// TIA Portal project "THELMA3_200224" (V15.1) (continued)
VERSION : 0.1
   STRUCT
      RemoteAddress : String;
      NonMDR_LabelName : String;
      "Date" : String;
      "Time" : String;
      RData : Array[0..56] of Byte;
      RdataBatch : Array[0..56] of Byte;
      BatchOK : Bool;
      TimeOK : Bool;
      AlarmCheck : Bool;
      LabelOK : Bool;
      LED_State : USInt;
      TimeDateError : Bool;
      Initialization : Bool;
      OPC_Error : Bool;
      TCP_ComError : Bool;
      TCP_ComErrorBatch : Bool;
      ComErrorStatus : Byte;
      ComErrorStatusBatch : Byte;
   END_STRUCT;
END_TYPE

TYPE "typeLCom_Config"
VERSION : 0.1
   STRUCT
      connection : Struct
         interfaceID : Hw_Any := 64;
         connectionID : Conn_Any := W#16#0FFF;
         comService : USInt := 2;
         isClient : Bool := false;
         localPort : UInt := 3456;
         partnerPort : UInt := 3456;
         partnerIP : IP_V4;
         acceptUnknownPartner : Bool := true;
         lifeSignCycleTime : Time := T#1s;
      END_STRUCT;
      sender : Struct
         cycleTime : Time := T#1s;
         ackTimeout : Time := T#1s;
      END_STRUCT;
      timeSync : Struct
         usePartnerTimestamps : Bool := false;
         sendMode : USInt;
         cycleTime : Time := T#1h;
         sendAtTimeOfDay : Time_Of_Day :=  TOD#05:00:0.000;
      END_STRUCT;
   END_STRUCT;
END_TYPE

TYPE "typeLCom_Diagnostics"
VERSION : 0.1
   STRUCT
      localConfig : Struct
         connection : Struct
            interfaceID : Hw_Any := 0;
            connectionID : Conn_Any := W#16#0000;
            comService : USInt := 0;
            isClient : Bool := false;
            localPort : UInt := 0;
            localIP : IP_V4;
            partnerPort : UInt := 3456;
            partnerIP : IP_V4;
            acceptUnknownPartner : Bool := false;
            useLComProtocol : Bool := false;
            lifeSignCycleTime : Time := T#0ms;
         END_STRUCT;
         sender : Struct
            cycleTime : Time;
            ackTimeout : Time;
         END_STRUCT;
         timeSync : Struct
            usePartnerTimestamps : Bool := false;
            sendMode : USInt;
            cycleTime : Time := T#0ms;
            sendAtTimeOfDay : Time_Of_Day :=  TOD#00:00:0.000;
         END_STRUCT;
         sizeOfSendBuffer : UDInt;
         sizeOfReceiveBuffer : UDInt;
      END_STRUCT;
      partnerConfig : Struct
         connnection : Struct
            lifeSignCycleTime : Time := T#0ms;
         END_STRUCT;
         sender : Struct
            cycleTime : Time := T#0ms;
            ackTimeout : Time := T#0ms;
         END_STRUCT;
         timeSync : Struct
            usePartnerTimestamps : Bool := false;
            sendMode : USInt;
         END_STRUCT;
         sizeOfSendBuffer : UDInt;
         sizeOfReceiveBuffer : UDInt;
      END_STRUCT;
      statistics : Struct
         avgCallCycle : Real;
         avgReceiveMsgCycle : Real;
         maxReceiveMsgCycle : Time;
         LComProtocolUsed : Bool := false;
         activeLComVersion : USInt;
         avgMsgSendingTime : Real;
         maxMsgSendingTime : Time;
         avgMsgReceivingTime : Real;
         maxMsgReceivingTime : Time;
         numberOfSentMessages : UDInt;
         numberOfReceivedMessages : UDInt;
         totalAckTimeouts : UInt;
         totalSendCycleViolations : UInt;
         totalReceiveCycleViolations : UInt;
         totalReconnects : UInt;
         lastConnect : DTL;
         lastTimeSync : DTL;
      END_STRUCT;
      bufferIndex : USInt := 16#FF;
      buffer : Array[0..63] of Struct
         status : Word;
         timestamp : DTL;
         isActive : Bool;
         subFunctionErrorID : Word;
         additionalValue1 : Real;
         additionalValue2 : Real;
         additionalValue3 : Real;
         additionalValue4 : Time;
      END_STRUCT;
   END_STRUCT;
   // buffer[1].isActive := false;
   // buffer[0].isActive := false;
   // buffer[2].isActive := false;
   // buffer[3].isActive := false;
   // buffer[4].isActive := false;
   // buffer[5].isActive := false;
   // buffer[6].isActive := false;
   // buffer[7].isActive := false;
   // buffer[8].isActive := false;
   // buffer[9].isActive := false;
   // buffer[10].isActive := false;
   // buffer[11].isActive := false;
   // buffer[12].isActive := false;
   // buffer[13].isActive := false;
   // buffer[14].isActive := false;
   // buffer[15].isActive := false;
   // buffer[16].isActive := false;
   // buffer[17].isActive := false;
   // buffer[18].isActive := false;
   // buffer[19].isActive := false;
   // buffer[20].isActive := false;
   // buffer[21].isActive := false;
   // buffer[22].isActive := false;
   // buffer[23].isActive := false;
   // buffer[24].isActive := false;
   // buffer[25].isActive := false;
   // buffer[26].isActive := false;
   // buffer[27].isActive := false;
   // buffer[28].isActive := false;
   // buffer[29].isActive := false;
   // buffer[30].isActive := false;
   // buffer[31].isActive := false;
   // buffer[32].isActive := false;
   // buffer[33].isActive := false;
   // buffer[34].isActive := false;
   // buffer[35].isActive := false;
   // buffer[36].isActive := false;
   // buffer[37].isActive := false;
   // buffer[38].isActive := false;
   // buffer[39].isActive := false;
   // buffer[40].isActive := false;
   // buffer[41].isActive := false;
   // buffer[42].isActive := false;
   // buffer[43].isActive := false;
   // buffer[44].isActive := false;
   // buffer[45].isActive := false;
   // buffer[46].isActive := false;
   // buffer[47].isActive := false;
   // buffer[48].isActive := false;
   // buffer[49].isActive := false;
   // buffer[50].isActive := false;
   // buffer[51].isActive := false;
   // buffer[52].isActive := false;
   // buffer[53].isActive := false;
   // buffer[54].isActive := false;
   // buffer[55].isActive := false;
   // buffer[56].isActive := false;
   // buffer[57].isActive := false;
   // buffer[58].isActive := false;
   // buffer[59].isActive := false;
   // buffer[60].isActive := false;
   // buffer[61].isActive := false;
   // buffer[62].isActive := false;
   // buffer[63].isActive := false;
END_TYPE

DATA_BLOCK "Skuska"   // DB1
{ S7_Optimized_Access := 'TRUE' }
VERSION : 0.1
   VAR
      SkuskaString : String;
      Length : Int;
      SkuskaArray : Array[0..56] of Byte;
      SkuskaString2 : String;
      TestBits : Array[0..10] of Bool;
      RemoteAdress : String := '192.168.1.10:29043';
   END_VAR
BEGIN
END_DATA_BLOCK

DATA_BLOCK "OPC"   // DB2
{ S7_Optimized_Access := 'TRUE' }
VERSION : 0.1
   VAR RETAIN
      CON_Material : "UDT_CON_Comm";
      TRP_Material : "UDT_TRP_Comm";
   END_VAR
BEGIN
END_DATA_BLOCK

DATA_BLOCK "SeP"   // DB3
{ S7_Optimized_Access := 'TRUE' }
VERSION : 0.1
   VAR
      Material_1 : "UDT_Status";
      Material_2 : "UDT_Status";
   END_VAR
BEGIN
END_DATA_BLOCK

DATA_BLOCK "LatestReading"   // DB4
{ S7_Optimized_Access := 'FALSE' }
VERSION : 0.1
   VAR
      TRP : "UDT_LatestReading";
   END_VAR
BEGIN
END_DATA_BLOCK

DATA_BLOCK "Reader"   // DB5
{ S7_Optimized_Access := 'TRUE' }
VERSION : 0.1
   VAR
      TRP : "UDT_Reader";
   END_VAR
BEGIN
END_DATA_BLOCK

DATA_BLOCK "TRP_DB"   // DB6
{ S7_Optimized_Access := 'TRUE' }
VERSION : 0.1
// stored: InstanceOfName TRP
"TRP"
BEGIN
END_DATA_BLOCK

DATA_BLOCK "CON_DB"   // DB7
{ S7_Optimized_Access := 'TRUE' }
VERSION : 0.1
// stored: InstanceOfName CON
"CON"
BEGIN
END_DATA_BLOCK

DATA_BLOCK "LatestReading_1"   // DB8
{ S7_Optimized_Access := 'FALSE' }
VERSION : 0.1
   VAR
      TRP : "UDT_LatestReading";
   END_VAR
BEGIN
END_DATA_BLOCK

DATA_BLOCK "PrinterData"   // DB9
{ S7_Optimized_Access := 'TRUE' }
VERSION : 0.1
   VAR RETAIN
      TRP : Struct
         PrinterData : "UDT_Printer";
         PrinterStatus : "typeLCom_Diagnostics";
         PrinterConfig : "typeLCom_Config";
      END_STRUCT;
      CON : Struct
         PrinterBagConfigBatch : "typeLCom_Config";
         PrinterBagStatusBatch : "typeLCom_Diagnostics";
         PrinterBagConfig : "typeLCom_Config";
         PrinterBagStatus : "typeLCom_Diagnostics";
         PrinterBagData : "UDT_CON_Printer";
         PrinterSelection : Bool;
      END_STRUCT;
   END_VAR
BEGIN
   TRP.PrinterData.RemoteAddress := '10.212.77.75:9100';
END_DATA_BLOCK

DATA_BLOCK "SiteCom"   // DB10
{ S7_Optimized_Access := 'FALSE' }
AUTHOR : nlagela
VERSION : 0.1
   VAR
      Material_1 : "UDT_ComMaterialReading";
      Material_2 : "UDT_ComMaterialReading";
   END_VAR
BEGIN
END_DATA_BLOCK

DATA_BLOCK "LatestReadings"   // DB11
{ S7_Optimized_Access := 'FALSE' }
VERSION : 0.1
   VAR
      Material_1 : "UDT_LatestReadingBag";
      Material_2 : "UDT_LatestReadingBag";
   END_VAR
BEGIN
END_DATA_BLOCK

DATA_BLOCK "PlainHandle_DB"   // DB12
{ S7_Optimized_Access := 'TRUE' }
VERSION : 0.1
// stored: InstanceOfName PlainHandle
"PlainHandle"
BEGIN
END_DATA_BLOCK

DATA_BLOCK "d10_PlainComm"   // DB13
{ S7_Optimized_Access := 'TRUE' }
VERSION : 0.1
   VAR
      Data_device : Array[0..7] of Bool;
   END_VAR
   VAR RETAIN
      bag_dmc_code : String [10];
      box_dmc_code : String [10];
      article_num : String [12];
      total_in_bag : String [7];
      total_in_box : String [7];
      product_weight : String [10];
      line_number : String [5];
      order_num : String [12];
   END_VAR
   VAR
      xPresetDataBagSent : Bool;
      xPresetDataBoxSent : Bool;
   END_VAR
BEGIN
END_DATA_BLOCK

DATA_BLOCK "d10_Data"   // DB14
{ S7_Optimized_Access := 'FALSE' }
VERSION : 0.1
   VAR
      Bag : Struct
         PlainCode : String[10];
         article_num : String[11];
         total_in_bag : String[6];
         total_in_box : String[6];
         product_weight : String[9];
         line_number : String[4];
         order_num : String[11];
         ReaderCode : Array[0..10] of Char;
      END_STRUCT;
      Box : Struct
         PlainCode : String[10];
         control1 : Bool;
      END_STRUCT;
      RawCode : String;
      Box_1 : Struct
         Box_Small_Code : String;
         Box_Code_1 : String[16];
         Box_Code_2 : String[12];
         Box_Code_3 : String[12];
         Box_Code_4 : String[16];
         Box_Code_5 : String[8];
         Box_Code_6 : String[8];
         Box_Code : String;
      END_STRUCT;
      Box_2 : Struct
         Box_Small_Code : String;
         Box_Code_1 : String[16];
         Box_Code_2 : String[12];
         Box_Code_3 : String[12];
         Box_Code_4 : String[16];
         Box_Code_5 : String[8];
         Box_Code_6 : String[8];
         Box_Code : String;
      END_STRUCT;
      Box_Codes : Struct
         Box_SmallCode : String[9];
         Box_LargeCode : String[80];
         Box_LargeCode_1 : String[16];
         Box_LargeCode_2 : String[12];
         Box_LargeCode_3 : String[12];
         Box_LargeCode_4 : String[16];
         Box_LargeCode_5 : String[8];
         Box_MIRAI_Code_6 : String[8];
      END_STRUCT;
      Code : String;
      RawArray : Array[0..86] of Char;
      TriggerDelayBag : Time;
      TriggerDelayBox : Time;
      NoEnigma : String := 'XXXXXXXXX';
      Empty : Array[0..79] of Char;
   END_VAR
BEGIN
END_DATA_BLOCK

DATA_BLOCK "d10_Alarms"   // DB15
{ S7_Optimized_Access := 'FALSE' }
AUTHOR : MCH
FAMILY : Fail
VERSION : 1.0
   VAR
      W_PLC : Struct
         "001" : Bool;
         "002" : Bool;
         "003" : Bool;
         "004" : Bool;
         "005" : Bool;
         "006" : Bool;
         "007" : Bool;
         "008" : Bool;
         "009" : Bool;
         "010" : Bool;
         "011" : Bool;
         "012" : Bool;
         "013" : Bool;
         "014" : Bool;
         "015" : Bool;
         "016" : Bool;
         "017" : Bool;
         "018" : Bool;
         "019" : Bool;
         "020" : Bool;
         "021" : Bool;
         "022" : Bool;
         "023" : Bool;
         "024" : Bool;
         "025" : Bool;
         "026" : Bool;
         "027" : Bool;
         "028" : Bool;
         "029" : Bool;
         "030" : Bool;
         "031" : Bool;
         "032" : Bool;
         "033" : Bool;
         "034" : Bool;
         "035" : Bool;
         "036" : Bool;
         "037" : Bool;
         "038" : Bool;
         "039" : Bool;
         "040" : Bool;
         "041" : Bool;
         "042" : Bool;
         "043" : Bool;
         "044" : Bool;
         "045" : Bool;
         "046" : Bool;
         "047" : Bool;
         "048" : Bool;
         "049" : Bool;
         "050" : Bool;
         "051" : Bool;
         "052" : Bool;
         "053" : Bool;
         "054" : Bool;
         "055" : Bool;
         "056" : Bool;
         "057" : Bool;
         "058" : Bool;
         "059" : Bool;
         "060" : Bool;
         "061" : Bool;
         "062" : Bool;
         "063" : Bool;
         "064" : Bool;
      END_STRUCT;
      W_HMI : Array[0..3] of Word;
      F_PLC : Struct
         "001" : Bool;
         "002" : Bool;
         "003" : Bool;
         "004" : Bool;
         "005" : Bool;
         "006" : Bool;
         "007" : Bool;
         "008" : Bool;
         "009" : Bool;
         "010" : Bool;
         "011" : Bool;
         "012" : Bool;
         "013" : Bool;
         "014" : Bool;
         "015" : Bool;
         "016" : Bool;
         "017" : Bool;
         "018" : Bool;
         "019" : Bool;
         "020" : Bool;
         "021" : Bool;
         "022" : Bool;
         "023" : Bool;
         "024" : Bool;
         "025" : Bool;
         "026" : Bool;
         "027" : Bool;
         "028" : Bool;
         "029" : Bool;
         "030" : Bool;
         "031" : Bool;
         "032" : Bool;
         "033" : Bool;
         "034" : Bool;
         "035" : Bool;
         "036" : Bool;
         "037" : Bool;
         "038" : Bool;
         "039" : Bool;
         "040" : Bool;
         "041" : Bool;
         "042" : Bool;
         "043" : Bool;
         "044" : Bool;
         "045" : Bool;
         "046" : Bool;
         "047" : Bool;
         "048" : Bool;
         "049" : Bool;
         "050" : Bool;
         "051" : Bool;
         "052" : Bool;
         "053" : Bool;
         "054" : Bool;
         "055" : Bool;
         "056" : Bool;
         "057" : Bool;
         "058" : Bool;
         "059" : Bool;
         "060" : Bool;
         "061" : Bool;
         "062" : Bool;
         "063" : Bool;
         "064" : Bool;
      END_STRUCT;
      F_HMI : Array[0..3] of Word;
   END_VAR
BEGIN
END_DATA_BLOCK

DATA_BLOCK "HMI"   // DB16
{ S7_Optimized_Access := 'TRUE' }
VERSION : 0.1
   VAR
      Control : Struct
         ResetFaults : Bool;
         NewRecipeLoaded : Bool;
         AutoRecipeFailed : Bool;
         RebootBag : Bool;
         RebootBox : Bool;
         Status : Int;
      END_STRUCT;
      Box_Small : Struct
         Control : Struct
            MaterialNumber : Bool;
            ResetCounters : Bool;
            TimeTrigger : Time;
            TcpCom : Bool;
         END_STRUCT;
         Codes : Struct
            MaterialNumberBox : UDInt;
            ActualReadingBox : UDInt;
         END_STRUCT;
         Counters : Struct
            CodeOk : DInt;
            CodeNok : DInt;
            CodeBadRead : DInt;
            Trigger : DInt;
            NewData : DInt;
            NDR : DInt;
         END_STRUCT;
      END_STRUCT;
      Box_Large : Struct
         Control : Struct
            MaterialNumber : Bool;
            ResetCounters : Bool;
            TimeTrigger : Time;
            TcpCom : Bool;
         END_STRUCT;
         Codes : Struct
            MaterialNumberBox : String;
            ActualReadingBox : String;
         END_STRUCT;
         Counters : Struct
            CodeOk : DInt;
            CodeNok : DInt;
            CodeBadRead : DInt;
            Trigger : DInt;
            NewData : DInt;
            NDR : DInt;
         END_STRUCT;
      END_STRUCT;
      Bag : Struct
         Control : Struct
            MaterialNumber : Bool;
            ResetCounters : Bool;
            TimeTrigger : Time;
            TcpCom : Bool;
         END_STRUCT;
         Codes : Struct
            MaterialNumberBox : UDInt;
            ActualReadingBox : UDInt;
         END_STRUCT;
         Counters : Struct
            CodeOk : DInt;
            CodeNok : DInt;
            CodeBadRead : DInt;
            Trigger : DInt;
            NewData : DInt;
            NDR : DInt;
         END_STRUCT;
      END_STRUCT;
   END_VAR
   VAR RETAIN
      Bag_Cam : Struct
         Vertiacal_position : Int;
         Horizontal_position : Int;
         Angle : Int;
         Delay_time_trigger : Int := 10;
         Fps : Int := 3;
      END_STRUCT;
      Box_Cam : Struct
         Vertiacal_position : Int;
         Horizontal_position : Int;
         Angle : Int;
         Delay_time_trigger : Int := 10;
         Fps : Int := 3;
      END_STRUCT;
   END_VAR
   VAR
      line_number_s : String;
      order_number_s : String;
      article_number_s : String;
      product_weight_s : String;
      total_in_bag_s : String;
      total_in_box_s : String;
      Enigma_off : Bool;
      Mirai_off : Bool;
   END_VAR
BEGIN
END_DATA_BLOCK

DATA_BLOCK "CodeHandle_DB"   // DB17
{ S7_Optimized_Access := 'TRUE' }
VERSION : 0.1
// stored: InstanceOfName CodeHandle
"CodeHandle"
BEGIN
END_DATA_BLOCK

DATA_BLOCK "DMCC_bag_DB"   // DB18
{ S7_Optimized_Access := 'TRUE' }
VERSION : 0.1
// stored: InstanceOfName DMCC_bag
"DMCC_bag"
BEGIN
END_DATA_BLOCK

DATA_BLOCK "ProgramReaderBox_IDB"   // DB21
{ S7_Optimized_Access := 'TRUE' }
VERSION : 0.1
// stored: InstanceOfName ProgramReaderBox
"ProgramReaderBox"
BEGIN
END_DATA_BLOCK

DATA_BLOCK "ProgramReaderBag_IDB"   // DB22
{ S7_Optimized_Access := 'TRUE' }
VERSION : 0.1
// stored: InstanceOfName ProgramReaderBag
"ProgramReaderBag"
BEGIN
END_DATA_BLOCK

DATA_BLOCK "d20_Alarms"   // DB25
{ S7_Optimized_Access := 'FALSE' }
AUTHOR : MCH
FAMILY : Fail
VERSION : 1.0
   VAR
      W_PLC : Struct
         "001" : Bool;
         "002" : Bool;
         "003" : Bool;
         "004" : Bool;
         "005" : Bool;
         "006" : Bool;
         "007" : Bool;
         "008" : Bool;
         "009" : Bool;
         "010" : Bool;
         "011" : Bool;
         "012" : Bool;
         "013" : Bool;
         "014" : Bool;
         "015" : Bool;
         "016" : Bool;
         "017" : Bool;
         "018" : Bool;
         "019" : Bool;
         "020" : Bool;
         "021" : Bool;
         "022" : Bool;
         "023" : Bool;
         "024" : Bool;
         "025" : Bool;
         "026" : Bool;
         "027" : Bool;
         "028" : Bool;
         "029" : Bool;
         "030" : Bool;
         "031" : Bool;
         "032" : Bool;
         "033" : Bool;
         "034" : Bool;
         "035" : Bool;
         "036" : Bool;
         "037" : Bool;
         "038" : Bool;
         "039" : Bool;
         "040" : Bool;
         "041" : Bool;
         "042" : Bool;
         "043" : Bool;
         "044" : Bool;
         "045" : Bool;
         "046" : Bool;
         "047" : Bool;
         "048" : Bool;
         "049" : Bool;
         "050" : Bool;
         "051" : Bool;
         "052" : Bool;
         "053" : Bool;
         "054" : Bool;
         "055" : Bool;
         "056" : Bool;
         "057" : Bool;
         "058" : Bool;
         "059" : Bool;
         "060" : Bool;
         "061" : Bool;
         "062" : Bool;
         "063" : Bool;
         "064" : Bool;
         "065" : Bool;
         "066" : Bool;
         "067" : Bool;
         "068" : Bool;
         "069" : Bool;
         "070" : Bool;
         "071" : Bool;
         "072" : Bool;
         "073" : Bool;
         "074" : Bool;
         "075" : Bool;
         "076" : Bool;
         "077" : Bool;
         "078" : Bool;
         "079" : Bool;
         "080" : Bool;
         "081" : Bool;
         "082" : Bool;
         "083" : Bool;
         "084" : Bool;
         "085" : Bool;
         "086" : Bool;
         "087" : Bool;
         "088" : Bool;
         "089" : Bool;
         "090" : Bool;
         "091" : Bool;
         "092" : Bool;
         "093" : Bool;
         "094" : Bool;
         "095" : Bool;
         "096" : Bool;
         "097" : Bool;
         "098" : Bool;
         "099" : Bool;
         "100" : Bool;
         "101" : Bool;
         "102" : Bool;
         "103" : Bool;
         "104" : Bool;
         "105" : Bool;
         "106" : Bool;
         "107" : Bool;
         "108" : Bool;
         "109" : Bool;
         "110" : Bool;
         "111" : Bool;
         "112" : Bool;
         "113" : Bool;
         "114" : Bool;
         "115" : Bool;
         "116" : Bool;
         "117" : Bool;
         "118" : Bool;
         "119" : Bool;
         "120" : Bool;
         "121" : Bool;
         "122" : Bool;
         "123" : Bool;
         "124" : Bool;
         "125" : Bool;
         "126" : Bool;
         "127" : Bool;
         "128" : Bool;
      END_STRUCT;
      W_HMI : Array[0..7] of Word;
      F_PLC : Struct
         "001" : Bool;
         "002" : Bool;
         "003" : Bool;
         "004" : Bool;
         "005" : Bool;
         "006" : Bool;
         "007" : Bool;
         "008" : Bool;
         "009" : Bool;
         "010" : Bool;
         "011" : Bool;
         "012" : Bool;
         "013" : Bool;
         "014" : Bool;
         "015" : Bool;
         "016" : Bool;
         "017" : Bool;
         "018" : Bool;
         "019" : Bool;
         "020" : Bool;
         "021" : Bool;
         "022" : Bool;
         "023" : Bool;
         "024" : Bool;
         "025" : Bool;
         "026" : Bool;
         "027" : Bool;
         "028" : Bool;
         "029" : Bool;
         "030" : Bool;
         "031" : Bool;
         "032" : Bool;
         "033" : Bool;
         "034" : Bool;
         "035" : Bool;
         "036" : Bool;
         "037" : Bool;
         "038" : Bool;
         "039" : Bool;
         "040" : Bool;
         "041" : Bool;
         "042" : Bool;
         "043" : Bool;
         "044" : Bool;
         "045" : Bool;
         "046" : Bool;
         "047" : Bool;
         "048" : Bool;
         "049" : Bool;
         "050" : Bool;
         "051" : Bool;
         "052" : Bool;
         "053" : Bool;
         "054" : Bool;
         "055" : Bool;
         "056" : Bool;
         "057" : Bool;
         "058" : Bool;
         "059" : Bool;
         "060" : Bool;
         "061" : Bool;
         "062" : Bool;
         "063" : Bool;
         "064" : Bool;
         "065" : Bool;
         "066" : Bool;
         "067" : Bool;
         "068" : Bool;
         "069" : Bool;
         "070" : Bool;
         "071" : Bool;
         "072" : Bool;
         "073" : Bool;
         "074" : Bool;
         "075" : Bool;
         "076" : Bool;
         "077" : Bool;
         "078" : Bool;
         "079" : Bool;
         "080" : Bool;
         "081" : Bool;
         "082" : Bool;
         "083" : Bool;
         "084" : Bool;
         "085" : Bool;
         "086" : Bool;
         "087" : Bool;
         "088" : Bool;
         "089" : Bool;
         "090" : Bool;
         "091" : Bool;
         "092" : Bool;
         "093" : Bool;
         "094" : Bool;
         "095" : Bool;
         "096" : Bool;
         "097" : Bool;
         "098" : Bool;
         "099" : Bool;
         "100" : Bool;
         "101" : Bool;
         "102" : Bool;
         "103" : Bool;
         "104" : Bool;
         "105" : Bool;
         "106" : Bool;
         "107" : Bool;
         "108" : Bool;
         "109" : Bool;
         "110" : Bool;
         "111" : Bool;
         "112" : Bool;
         "113" : Bool;
         "114" : Bool;
         "115" : Bool;
         "116" : Bool;
         "117" : Bool;
         "118" : Bool;
         "119" : Bool;
         "120" : Bool;
         "121" : Bool;
         "122" : Bool;
         "123" : Bool;
         "124" : Bool;
         "125" : Bool;
         "126" : Bool;
         "127" : Bool;
         "128" : Bool;
      END_STRUCT;
      F_HMI : Array[0..15] of Word;
   END_VAR
BEGIN
END_DATA_BLOCK

DATA_BLOCK "X_Simulacia_DB"   // DB100
{ S7_Optimized_Access := 'TRUE' }
VERSION : 0.1
// stored: InstanceOfName X_Simulacia
"X_Simulacia"
BEGIN
   OPC_Con.NewMDR_Flag := '0123';
   OPC_Con.NewArticleFlag := '5987';
   OPC_Con.NewBatchNumber := '123456';
   OPC_Con.NewArtBaseNumber := 15478;
   OPC_Con.NewExtDate := '031219';
   OPC_Con.NewBatchEndTime := '103258';
   OPC_Con.NewMarketREG_Code := '879654';
END_DATA_BLOCK

DATA_BLOCK "DB_DMCC_Data"   // DB110
{ S7_Optimized_Access := 'FALSE' }
VERSION : 0.1
   VAR
      ResetChars_Camera_Box : Array[0..63] of Char;
      SetChars_Camera_Box : Array[0..63] of Char;
      ClearLogChars_Camera_Box : Array[0..63] of Char;
      ResetChars_Camera_Bag : Array[0..63] of Char;
      SetChars_Camera_Bag : Array[0..63] of Char;
      ClearLogChars_Camera_Bag : Array[0..63] of Char;
      Reboot_Box : Array[0..63] of Char;
      Reboot_Bag : Array[0..63] of Char;
   END_VAR
BEGIN
END_DATA_BLOCK

DATA_BLOCK "DMCC_DB_1"   // DB111
{ S7_Optimized_Access := 'TRUE' }
VERSION : 0.1
// stored: InstanceOfName DMCC
"DMCC"
BEGIN
END_DATA_BLOCK

FUNCTION_BLOCK "VideoJet_1520"   // FB1, FBD
{ S7_Optimized_Access := 'TRUE' }
VERSION : 0.1
   VAR_INPUT
      RemoteAddress : String[20] := '10.176.40.90';
      ConnectionStatus : Bool;
      ID : Conn_Ouc;
      ConType : Bool;
      ArtFlag : Bool;
      MDR_Flag : Bool;
      BatchStatus : USInt;
      BatchNumber : String;
      ArtBaseNumber : String;
      MarketRegCode : String;
      ExtDate : String;
      PlainDataChanged : Bool;
      "Date" : String;
      "Time" : String;
      DataReceived : Bool;
      DataSent : Bool;
      TimeSynchPeriod : Time := T#10M;
      AlarmCheckPeriod : Time := T#5M;
      RData : Array[0..56] of Byte;
      NMDR_LabelName : String;
      LabelSelecting : Bool;
   END_VAR
   VAR_OUTPUT
      ErrorIP : Bool;
      BatchOK : Bool;
      AlarmCheck : Bool;
      TimeOK : Bool;
      LabelOK : Bool;
   END_VAR
   VAR
      Config : TADDR_Param;
      Configuration : "typeLCom_Config";
      RLen : UDInt;
      SLen : UDInt;
      SData : Array[0..56] of Byte;
      StartTNR : Bool;
      TimeNR : Time := T#1m;
      SendAgainTrigger : Bool;
      NotReceiveT : TON_TIME;
      TimeSynchEnable : Bool := false;
      TimeSynchT : TON_TIME;
      AlarmCheckEnable : Bool := false;
      AlarmCheckT : TON_TIME;
      STrig : Bool;
      "Step" : UDInt;
      AlarmReceivedData : Array[0..56] of Byte;
      PrinterAlarmStatus : Array[0..8] of Char;
      TimeReceivedData : Array[0..56] of Byte;
      BatchReceivedData : Array[0..56] of Byte;
      BBD_ReceivedData : Array[0..56] of Byte;
      LabelReceivedData : Array[0..56] of Byte;
      RdataTime : Bool;
      RdataAlarm : Bool;
      RdataBatch : Bool;
      RdataBBD : Bool;
      RdataLabel : Bool;
      BlockedProduct : Bool;
      DateChar : Array[0..7] of Char;
      ReconnectR : R_TRIG;
      MDR_R : R_TRIG;
      MDR_F : F_TRIG;
      BlockedR : R_TRIG;
      BlockedF : F_TRIG;
      ActualNMDR_Label : String;
      NLabelChanged : Bool;
      Selected : Bool;
      First : Bool;
      SelectingR : R_TRIG;
      BatchAfterLabelT : TON_TIME;
      SecondAfterFirstT : TON_TIME;
      BBD_OK : Bool;
      ChangeIP_T : TP_TIME;
      IP_Change : Bool;
      RemoteAddressOld : String;
   END_VAR
   VAR_TEMP
      StatusIP : Word;
      Dummy2 : UInt;
      i : Int;
      CommandHead : String;
      BatchNumSTR : String;
      BatchNumberChar : Array[0..10] of Char;
      SDataDummy : String;
      LenDummy : Int;
      LenLabel : Int;
      DateDummy : String;
   END_VAR
   VAR CONSTANT
      Start : Char := '$02';
      End : Char := '$03';
      NewLine : Char := '$L';
      FirstField : String := 'BATCH_ART';
      SecondField : String := 'MARKE_BBD';
      MDR_LabelName : String := 'MDR';
   END_VAR
BEGIN

REGION Network 1 (SCL)
   //---------------------------------------------------------------------
   //In this network first, we assign the ip address and port number for the printer (VideoJet). Then prepare the command for 
   //time synch, receiving alarms, sending a batch number and selectiong the label. one port for all data.
   //---------------------------------------------------------------------
   //
   REGION Address_Assign
       (*
       //Special case: if ip and port is entered correctly but still the communication not established, try onece more.
       IF #ConnectionStatus = False AND #ErrorIP = FALSE AND #ReTry = FALSE AND #ConnAgainT.Q = FALSE AND #TimeOutError = FALSE THEN
           #ReTry := True;
       ELSE
           #ReTry := FALSE;
       END_IF;
       *)
       // ip and port assign to the printer
       #Config := "LGF_StringToTaddr"(ipAddressString := #RemoteAddress, error => #ErrorIP, status => #StatusIP);
       //when IP address change, disconnect and connect again
       #ChangeIP_T(IN := #RemoteAddressOld <> #RemoteAddress,
                   PT := T#2S);
       IF #ChangeIP_T.Q OR #ErrorIP = TRUE THEN
           #IP_Change := TRUE;
       ELSE
           #IP_Change := FALSE;
       END_IF;
       #RemoteAddressOld := #RemoteAddress;
       FOR #i := 1 TO 4 DO
           #Configuration.connection.partnerIP.ADDR[#i] := USINT_TO_BYTE(#Config.REM_IP_ADDR[#i]);//assign ip address
       END_FOR;
       //assign id port and other setting for TCP communication
       #Configuration.connection.connectionID := #ID;
       #Configuration.connection.comService := 1;
       //if it is active connection
       IF #ConType = TRUE THEN
           #Configuration.connection.isClient := True;
           IF #Config.REM_PORT_NR = 0 THEN
               #Configuration.connection.partnerPort :=3100; // default port for video jet communication
           ELSE
               #Configuration.connection.partnerPort := #Config.REM_PORT_NR;
           END_IF;
       ELSE //if it is passive connection
           #Configuration.connection.isClient := FALSE;
           #Configuration.connection.localPort := 2000;
       END_IF;
   END_REGION
   REGION Trigger
       // Trigger signal to send a correct data for print when Batch ended
       IF #BatchStatus = 3 THEN
           #BlockedProduct := TRUE;
       ELSE
           #BlockedProduct := FALSE;
       END_IF;
       // Trigger signal to send Non-MDR label when it is changed from the screen
       IF #MDR_Flag = FALSE AND #ActualNMDR_Label <> #NMDR_LabelName THEN
           #NLabelChanged := TRUE;
           #ActualNMDR_Label := #NMDR_LabelName;
       ELSE
           #NLabelChanged := FALSE;
       END_IF;
   END_REGION
   REGION Commands 
       // Creating Commands and preparing them to Send
       IF #Step = 1 THEN
           //command for time synchronisation
           #CommandHead := 'Z'; //head for time/date synch
           #SData[0] := #Start;
           Strg_TO_Chars(Strg := #CommandHead,
                         pChars := 1,
                         Cnt => #Dummy2,
                         Chars := #SData);
           #DateDummy := DELETE(IN := #Date, L := 2, P := 1);
           Strg_TO_Chars(Strg := #DateDummy,
                         pChars := 2,
                         Cnt => #Dummy2,
                         Chars := #SData);
           Strg_TO_Chars(Strg := #Time,
                         pChars := 8,
                         Cnt => #Dummy2,
                         Chars := #SData);
           #SData[14] := #End;
           #RLen := 3;
           #SLen := 15;
           #STrig := TRUE;
           #Step := 0; //idea state
           #RdataTime := TRUE;
           #RdataAlarm := FALSE;
           #RdataBatch := FALSE;
           #RdataBBD := FALSE;
           #RdataLabel := FALSE;
       ELSIF #Step = 2 THEN
           //command for checking the alarms
           #CommandHead := 'E'; //head for current status of the printer
           #SData[0] := #Start;
           Strg_TO_Chars(Strg := #CommandHead,
                         pChars := 1,
                         Cnt => #Dummy2,
                         Chars := #SData);
           #SData[2] := #End;
           #RLen := 9;
           #SLen := 3;
           #STrig := TRUE;
           #Step := 0;
           #RdataAlarm := TRUE;
           #RdataTime := FALSE;
           #RdataBatch := FALSE;
           #RdataBBD := FALSE;
           #RdataLabel := FALSE;
       ELSIF #Step = 3 THEN
           (*update first external field (batch and art number)
            You need TO create two seperate external fields with the name OF "BATCH_ART" AND "MARKET_BBD"*)
           #CommandHead := 'U'; //head for update user field
           #RLen := 3;
           #Step := 0;
           #STrig := TRUE;
           #RdataTime := FALSE;
           #RdataAlarm := FALSE;
           #RdataBatch := TRUE;
           #RdataBBD := FALSE;
           #RdataLabel := FALSE;
           #Selected := FALSE;
           #SData[0] := #Start;
           Strg_TO_Chars(Strg := #CommandHead,
                         pChars := 1,
                         Cnt => #Dummy2,
                         Chars := #SData);
           #SDataDummy := CONCAT(IN1 := #FirstField, IN2 := #NewLine);
           Strg_TO_Chars(Strg := #SDataDummy,
                         pChars := 2,
                         Cnt => #Dummy2,
                         Chars := #SData);
           IF #ArtFlag = TRUE THEN
               #LenDummy := LEN(#ArtBaseNumber);
               #SDataDummy := CONCAT(IN1 := #BatchNumber, IN2 := ' ');
               #SDataDummy := CONCAT(IN1 := #SDataDummy, IN2 := 'ART');
               #SDataDummy := CONCAT(IN1 := #SDataDummy, IN2 := #ArtBaseNumber);
               IF #BatchStatus = 3 THEN //add a sign '+' at the con
                   #SDataDummy := CONCAT(IN1 := #SDataDummy, IN2 := '+');
               ELSE
                   #SDataDummy := CONCAT(IN1 := #SDataDummy, IN2 := ' ');
               END_IF;
               Strg_TO_Chars(Strg := #SDataDummy,
                             pChars := 12,
                             Cnt => #Dummy2,
                             Chars := #SData);
               #SData[15 + 12 + #LenDummy] := #End;
               #SLen := 15 + 12 + #LenDummy + 1;
           ELSE //no print article number
               IF #BatchStatus = 3 THEN //add a sign '+' at the con
                   #SDataDummy := CONCAT(IN1 := #BatchNumber, IN2 := '+');
               ELSE
                   #SDataDummy := CONCAT(IN1 := #BatchNumber, IN2 := ' ');
               END_IF;
               Strg_TO_Chars(Strg := #SDataDummy,
                             pChars := 12,
                             Cnt => #Dummy2,
                             Chars := #SData);
               #SData[23] := #End;
               #SLen := 24;
           END_IF;
       ELSIF #Step = 4 THEN
           (*update second external field (batch and art number)
                  You need TO create two seperate external fields with the name OF "BATCH_ART" AND "MARKE_BBD"*)
           #SData[0] := #Start;
           #First := FALSE;
           IF #MarketRegCode = '' AND #ExtDate = '' THEN // delete second row data
               #CommandHead := 'D'; //head for update user field
               #SDataDummy := CONCAT(IN1 := #CommandHead, IN2 := #SecondField);
               Strg_TO_Chars(Strg := #SDataDummy,
                             pChars := 1,
                             Cnt => #Dummy2,
                             Chars := #SData);
               #SData[11] := #End;
               #SLen := 12;
               #RLen := 3;
               #Step := 0;
               #STrig := TRUE;
               #RdataTime := FALSE;
               #RdataAlarm := FALSE;
               #RdataBatch := FALSE;
               #RdataBBD := TRUE;
               #RdataLabel := FALSE;
               #Selected := FALSE;
           ELSIF #MarketRegCode <> '' AND #ExtDate = '' THEN // only print market reg code on the second row
               #CommandHead := 'U'; //head for update user field
               #LenDummy := LEN(#MarketRegCode);
               #SDataDummy := CONCAT(IN1 := #CommandHead, IN2 := #SecondField);
               #SDataDummy := CONCAT(IN1 := #SDataDummy, IN2 := #NewLine);
               #SDataDummy := CONCAT(IN1 := #SDataDummy, IN2 := #MarketRegCode);
               Strg_TO_Chars(Strg := #SDataDummy,
                             pChars := 1,
                             Cnt => #Dummy2,
                             Chars := #SData);
               #SData[12 + #LenDummy] := #End;
               #SLen := 12 + #LenDummy + 1;
               #RLen := 3;
               #Step := 0;
               #STrig := TRUE;
               #RdataTime := FALSE;
               #RdataAlarm := FALSE;
               #RdataBatch := FALSE;
               #RdataBBD := TRUE;
               #RdataLabel := FALSE;
               #Selected := FALSE;
           ELSIF #MarketRegCode = '' AND #ExtDate <> '' THEN // only print best before date on the second row
               #CommandHead := 'U'; //head for update user field
               #LenDummy := LEN(#ExtDate);
               #SDataDummy := CONCAT(IN1 := #CommandHead, IN2 := #SecondField);
               #SDataDummy := CONCAT(IN1 := #SDataDummy, IN2 := #NewLine);